                           Sts_FilterExcludedNumEvents => #instEventSortFilter_Alarm.Sts_FilterExcludedNumEvents,
                           Sts_SortFilterNumEvents => #instEventSortFilter_Alarm.Sts_SortFilterNumEvents);
END_REGION

REGION Network 10: *** Beging the WARNING area ****
END_REGION

REGION Network 11: Warning Event Summary Logic - Beginning Block
   // **********  WARNING SUMMATION  **********
   //  
   // The event summation begin instruction prepares the summation blocks.  It should be run each time before the FB_EventSummation blocks.
   RUNG wire#powerrail
      #instEventSumBeg_Warning(Sts_EventSummation := "Warning".Summation)
   END_RUNG
   // the same network as SCL:
   #instEventSumBeg_Warning(Sts_EventSummation := "Warning".Summation);   // "CPG_EventSummationBegin"
END_REGION

REGION Network 12: Warning Event Summary Logic - Unit Level Warnings
   RUNG wire#powerrail
      Contact( "UN".PackML_Sts.moduleActive )
      I_Contact( "HMI_Data".EMSortDisableWarning.Unit )
      #instEventSum_Warning_UN(In_EventStatus := "UN".Warning, Sts_EventSummation := "Warning".Summation, Sts_NumEvents => #instEventSum_Warning_UN.Sts_NumEvents, Sts_Category_0_Latched =>, Sts_Category_1_Latched =>, Sts_Category_2_Latched =>, Sts_Category_3_Latched =>, Sts_Category_4_Latched =>, Sts_Category_5_Latched =>, Sts_Category_6_Latched =>, Sts_Category_7_Latched =>, Sts_Category_8_Latched =>, Sts_Category_9_Latched =>, Sts_Category_0_NotLatched =>, Sts_Category_1_NotLatched =>, Sts_Category_2_NotLatched =>, Sts_Category_3_NotLatched =>, Sts_Category_4_NotLatched =>, Sts_Category_5_NotLatched =>, Sts_Category_6_NotLatched =>, Sts_Category_7_NotLatched =>, Sts_Category_8_NotLatched =>, Sts_Category_9_NotLatched =>, Sts_CurrentActiveEvent => #instEventSum_Warning_UN.Sts_CurrentActiveEvent, Sts_Error => #instEventSum_Warning_UN.Sts_Error, Sts_ErrorCode => #instEventSum_Warning_UN.Sts_ErrorCode)
   END_RUNG
   // the same network as SCL:
   IF "UN".PackML_Sts.moduleActive AND NOT "HMI_Data".EMSortDisableWarning.Unit THEN
       #instEventSum_Warning_UN(In_EventStatus := "UN".Warning,   // "CPG_EventSummation"
                               Sts_EventSummation := "Warning".Summation,
                               Sts_NumEvents => #instEventSum_Warning_UN.Sts_NumEvents,
                               Sts_CurrentActiveEvent => #instEventSum_Warning_UN.Sts_CurrentActiveEvent,
                               Sts_Error => #instEventSum_Warning_UN.Sts_Error,
                               Sts_ErrorCode => #instEventSum_Warning_UN.Sts_ErrorCode);
   END_IF;
END_REGION

REGION Network 13: Warning Event Summary Logic - Equipment Module #00
   // This instance of the Event Sum (or Event Summation) is used to merge the events 
   // from EM0 into the larger Unit or UN evevts list.
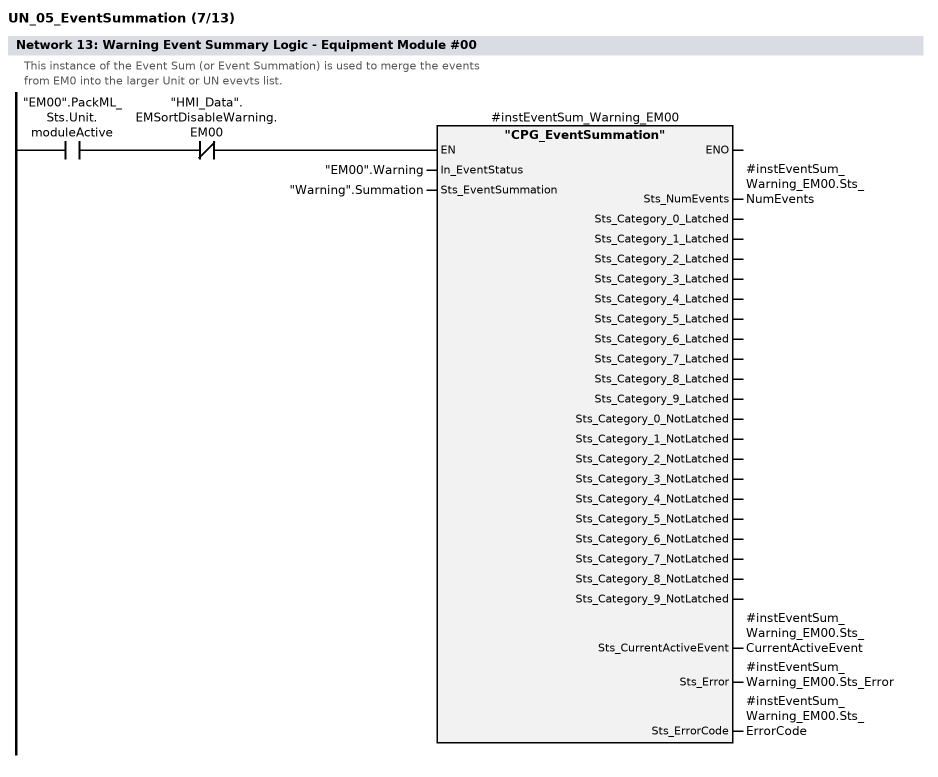
   RUNG wire#powerrail
      Contact( "EM00".PackML_Sts.Unit.moduleActive )
      I_Contact( "HMI_Data".EMSortDisableWarning.EM00 )
      #instEventSum_Warning_EM00(In_EventStatus := "EM00".Warning, Sts_EventSummation := "Warning".Summation, Sts_NumEvents => #instEventSum_Warning_EM00.Sts_NumEvents, Sts_Category_0_Latched =>, Sts_Category_1_Latched =>, Sts_Category_2_Latched =>, Sts_Category_3_Latched =>, Sts_Category_4_Latched =>, Sts_Category_5_Latched =>, Sts_Category_6_Latched =>, Sts_Category_7_Latched =>, Sts_Category_8_Latched =>, Sts_Category_9_Latched =>, Sts_Category_0_NotLatched =>, Sts_Category_1_NotLatched =>, Sts_Category_2_NotLatched =>, Sts_Category_3_NotLatched =>, Sts_Category_4_NotLatched =>, Sts_Category_5_NotLatched =>, Sts_Category_6_NotLatched =>, Sts_Category_7_NotLatched =>, Sts_Category_8_NotLatched =>, Sts_Category_9_NotLatched =>, Sts_CurrentActiveEvent => #instEventSum_Warning_EM00.Sts_CurrentActiveEvent, Sts_Error => #instEventSum_Warning_EM00.Sts_Error, Sts_ErrorCode => #instEventSum_Warning_EM00.Sts_ErrorCode)
   END_RUNG
   // the same network as SCL:
   IF "EM00".PackML_Sts.Unit.moduleActive AND NOT "HMI_Data".EMSortDisableWarning.EM00 THEN
       #instEventSum_Warning_EM00(In_EventStatus := "EM00".Warning,   // "CPG_EventSummation"
                               Sts_EventSummation := "Warning".Summation,
                               Sts_NumEvents => #instEventSum_Warning_EM00.Sts_NumEvents,
                               Sts_CurrentActiveEvent => #instEventSum_Warning_EM00.Sts_CurrentActiveEvent,
                               Sts_Error => #instEventSum_Warning_EM00.Sts_Error,
                               Sts_ErrorCode => #instEventSum_Warning_EM00.Sts_ErrorCode);
   END_IF;
END_REGION

REGION Network 14: Warning Event Summary Logic - Equipment Module #01
   // This instance of the Event Sum (or Event Summation) is used to merge the events 
   // from EM1 into the larger Unit or UN evevts list.
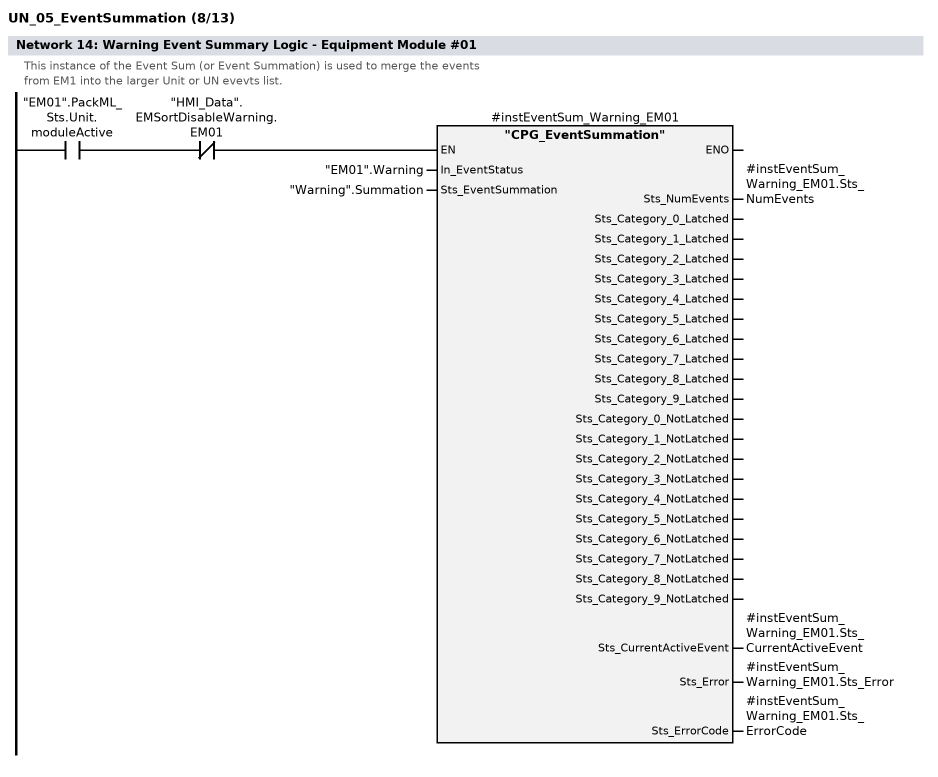
   RUNG wire#powerrail
      Contact( "EM01".PackML_Sts.Unit.moduleActive )
      I_Contact( "HMI_Data".EMSortDisableWarning.EM01 )
      #instEventSum_Warning_EM01(In_EventStatus := "EM01".Warning, Sts_EventSummation := "Warning".Summation, Sts_NumEvents => #instEventSum_Warning_EM01.Sts_NumEvents, Sts_Category_0_Latched =>, Sts_Category_1_Latched =>, Sts_Category_2_Latched =>, Sts_Category_3_Latched =>, Sts_Category_4_Latched =>, Sts_Category_5_Latched =>, Sts_Category_6_Latched =>, Sts_Category_7_Latched =>, Sts_Category_8_Latched =>, Sts_Category_9_Latched =>, Sts_Category_0_NotLatched =>, Sts_Category_1_NotLatched =>, Sts_Category_2_NotLatched =>, Sts_Category_3_NotLatched =>, Sts_Category_4_NotLatched =>, Sts_Category_5_NotLatched =>, Sts_Category_6_NotLatched =>, Sts_Category_7_NotLatched =>, Sts_Category_8_NotLatched =>, Sts_Category_9_NotLatched =>, Sts_CurrentActiveEvent => #instEventSum_Warning_EM01.Sts_CurrentActiveEvent, Sts_Error => #instEventSum_Warning_EM01.Sts_Error, Sts_ErrorCode => #instEventSum_Warning_EM01.Sts_ErrorCode)
   END_RUNG
   // the same network as SCL:
   IF "EM01".PackML_Sts.Unit.moduleActive AND NOT "HMI_Data".EMSortDisableWarning.EM01 THEN
       #instEventSum_Warning_EM01(In_EventStatus := "EM01".Warning,   // "CPG_EventSummation"
                               Sts_EventSummation := "Warning".Summation,
                               Sts_NumEvents => #instEventSum_Warning_EM01.Sts_NumEvents,
                               Sts_CurrentActiveEvent => #instEventSum_Warning_EM01.Sts_CurrentActiveEvent,
                               Sts_Error => #instEventSum_Warning_EM01.Sts_Error,
                               Sts_ErrorCode => #instEventSum_Warning_EM01.Sts_ErrorCode);
   END_IF;
END_REGION

REGION Network 15: Warning Event Summary Logic - Equipment Module #02
   // This instance of the Event Sum (or Event Summation) is used to merge the events 
   // from EM01 into the larger Unit or UN evevts list.
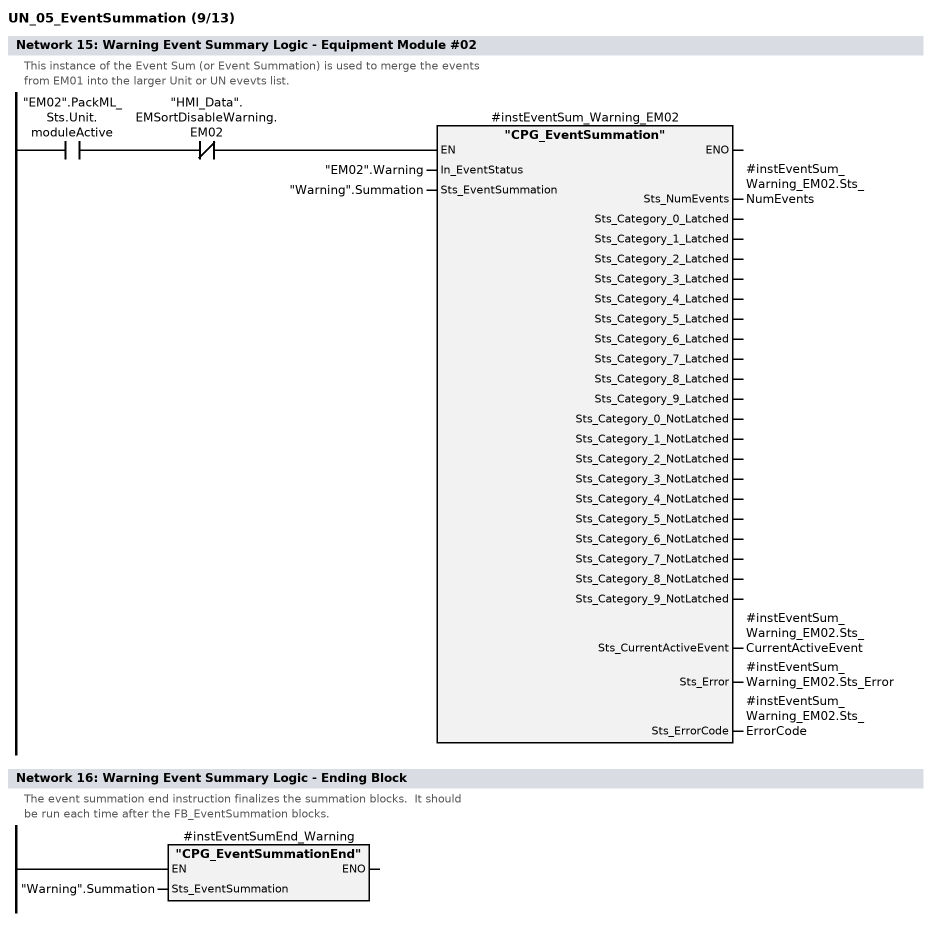
   RUNG wire#powerrail
      Contact( "EM02".PackML_Sts.Unit.moduleActive )
      I_Contact( "HMI_Data".EMSortDisableWarning.EM02 )
      #instEventSum_Warning_EM02(In_EventStatus := "EM02".Warning, Sts_EventSummation := "Warning".Summation, Sts_NumEvents => #instEventSum_Warning_EM02.Sts_NumEvents, Sts_Category_0_Latched =>, Sts_Category_1_Latched =>, Sts_Category_2_Latched =>, Sts_Category_3_Latched =>, Sts_Category_4_Latched =>, Sts_Category_5_Latched =>, Sts_Category_6_Latched =>, Sts_Category_7_Latched =>, Sts_Category_8_Latched =>, Sts_Category_9_Latched =>, Sts_Category_0_NotLatched =>, Sts_Category_1_NotLatched =>, Sts_Category_2_NotLatched =>, Sts_Category_3_NotLatched =>, Sts_Category_4_NotLatched =>, Sts_Category_5_NotLatched =>, Sts_Category_6_NotLatched =>, Sts_Category_7_NotLatched =>, Sts_Category_8_NotLatched =>, Sts_Category_9_NotLatched =>, Sts_CurrentActiveEvent => #instEventSum_Warning_EM02.Sts_CurrentActiveEvent, Sts_Error => #instEventSum_Warning_EM02.Sts_Error, Sts_ErrorCode => #instEventSum_Warning_EM02.Sts_ErrorCode)
   END_RUNG
   // the same network as SCL:
   IF "EM02".PackML_Sts.Unit.moduleActive AND NOT "HMI_Data".EMSortDisableWarning.EM02 THEN
       #instEventSum_Warning_EM02(In_EventStatus := "EM02".Warning,   // "CPG_EventSummation"
                               Sts_EventSummation := "Warning".Summation,
                               Sts_NumEvents => #instEventSum_Warning_EM02.Sts_NumEvents,
                               Sts_CurrentActiveEvent => #instEventSum_Warning_EM02.Sts_CurrentActiveEvent,
                               Sts_Error => #instEventSum_Warning_EM02.Sts_Error,
                               Sts_ErrorCode => #instEventSum_Warning_EM02.Sts_ErrorCode);
   END_IF;
END_REGION

REGION Network 16: Warning Event Summary Logic - Ending Block
   // The event summation end instruction finalizes the summation blocks.  It should 
   // be run each time after the FB_EventSummation blocks.
   RUNG wire#powerrail
      #instEventSumEnd_Warning(Sts_EventSummation := "Warning".Summation)
   END_RUNG
   // the same network as SCL:
   #instEventSumEnd_Warning(Sts_EventSummation := "Warning".Summation);   // "CPG_EventSummationEnd"
END_REGION

REGION Network 17: Event Sort Filter logic - Warnings
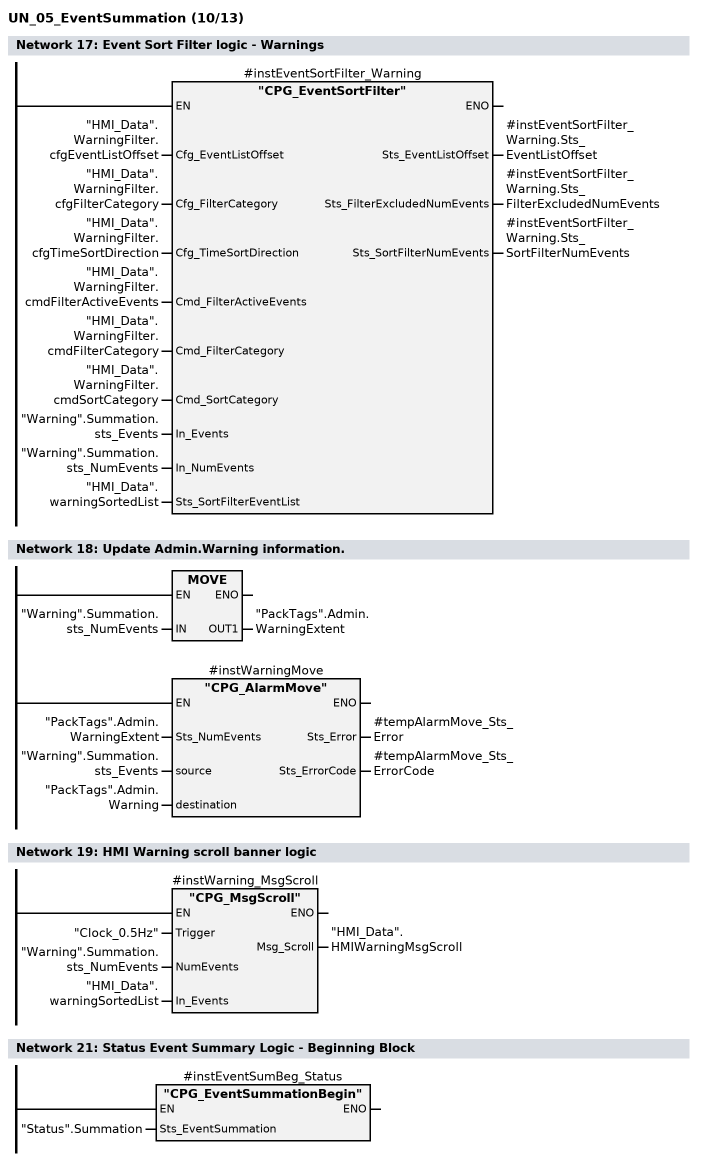
   RUNG wire#powerrail
      #instEventSortFilter_Warning(Cfg_EventListOffset := "HMI_Data".WarningFilter.cfgEventListOffset, Cfg_FilterCategory := "HMI_Data".WarningFilter.cfgFilterCategory, Cfg_TimeSortDirection := "HMI_Data".WarningFilter.cfgTimeSortDirection, Cmd_FilterActiveEvents := "HMI_Data".WarningFilter.cmdFilterActiveEvents, Cmd_FilterCategory := "HMI_Data".WarningFilter.cmdFilterCategory, Cmd_SortCategory := "HMI_Data".WarningFilter.cmdSortCategory, In_Events := "Warning".Summation.sts_Events, In_NumEvents := "Warning".Summation.sts_NumEvents, Sts_SortFilterEventList := "HMI_Data".warningSortedList, Sts_EventListOffset => #instEventSortFilter_Warning.Sts_EventListOffset, Sts_FilterExcludedNumEvents => #instEventSortFilter_Warning.Sts_FilterExcludedNumEvents, Sts_SortFilterNumEvents => #instEventSortFilter_Warning.Sts_SortFilterNumEvents)
   END_RUNG
   // the same network as SCL:
   #instEventSortFilter_Warning(Cfg_EventListOffset := "HMI_Data".WarningFilter.cfgEventListOffset,   // "CPG_EventSortFilter"
                           Cfg_FilterCategory := "HMI_Data".WarningFilter.cfgFilterCategory,
                           Cfg_TimeSortDirection := "HMI_Data".WarningFilter.cfgTimeSortDirection,
                           Cmd_FilterActiveEvents := "HMI_Data".WarningFilter.cmdFilterActiveEvents,
                           Cmd_FilterCategory := "HMI_Data".WarningFilter.cmdFilterCategory,
                           Cmd_SortCategory := "HMI_Data".WarningFilter.cmdSortCategory,
                           In_Events := "Warning".Summation.sts_Events,
                           In_NumEvents := "Warning".Summation.sts_NumEvents,
                           Sts_SortFilterEventList := "HMI_Data".warningSortedList,
                           Sts_EventListOffset => #instEventSortFilter_Warning.Sts_EventListOffset,
                           Sts_FilterExcludedNumEvents => #instEventSortFilter_Warning.Sts_FilterExcludedNumEvents,
                           Sts_SortFilterNumEvents => #instEventSortFilter_Warning.Sts_SortFilterNumEvents);
END_REGION

REGION Network 18: Update Admin.Warning information.
   RUNG wire#powerrail
      { S7_GenerateENO := "TRUE" } Move(in := "Warning".Summation.sts_NumEvents, out1 => "PackTags".Admin.WarningExtent)
   END_RUNG
   RUNG wire#powerrail
      #instWarningMove(Sts_NumEvents := "PackTags".Admin.WarningExtent, source := "Warning".Summation.sts_Events, destination := "PackTags".Admin.Warning, Sts_Error => #tempAlarmMove_Sts_Error, Sts_ErrorCode => #tempAlarmMove_Sts_ErrorCode)
   END_RUNG
   // the same network as SCL:
   "PackTags".Admin.WarningExtent := "Warning".Summation.sts_NumEvents;
   #instWarningMove(Sts_NumEvents := "PackTags".Admin.WarningExtent,   // "CPG_AlarmMove"
                    source := "Warning".Summation.sts_Events,
                    destination := "PackTags".Admin.Warning,
                    Sts_Error => #tempAlarmMove_Sts_Error,
                    Sts_ErrorCode => #tempAlarmMove_Sts_ErrorCode);
END_REGION

REGION Network 19: HMI Warning scroll banner logic
   RUNG wire#powerrail
      #instWarning_MsgScroll(Trigger := "Clock_0.5Hz", NumEvents := "Warning".Summation.sts_NumEvents, In_Events := "HMI_Data".warningSortedList, Msg_Scroll => "HMI_Data".HMIWarningMsgScroll)
   END_RUNG
   // the same network as SCL:
   #instWarning_MsgScroll(Trigger := "Clock_0.5Hz",   // "CPG_MsgScroll"
                          NumEvents := "Warning".Summation.sts_NumEvents,
                          In_Events := "HMI_Data".warningSortedList,
                          Msg_Scroll => "HMI_Data".HMIWarningMsgScroll);
END_REGION

REGION Network 20: *** Status Event Summation ***
END_REGION

REGION Network 21: Status Event Summary Logic - Beginning Block
   RUNG wire#powerrail
      #instEventSumBeg_Status(Sts_EventSummation := "Status".Summation)
   END_RUNG
   // the same network as SCL:
   #instEventSumBeg_Status(Sts_EventSummation := "Status".Summation);   // "CPG_EventSummationBegin"
END_REGION

REGION Network 22: Status Event Summary Logic - Unit
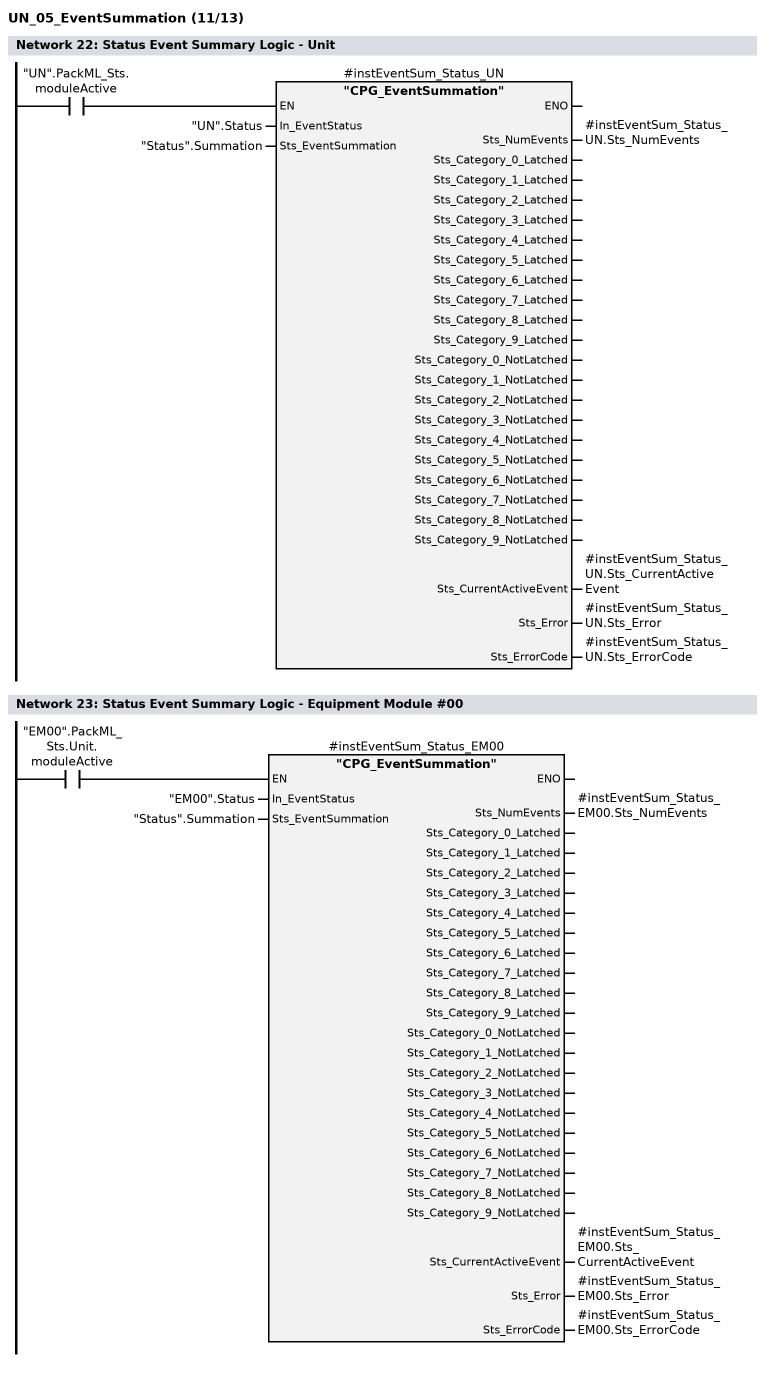
   RUNG wire#powerrail
      Contact( "UN".PackML_Sts.moduleActive )
      #instEventSum_Status_UN(In_EventStatus := "UN".Status, Sts_EventSummation := "Status".Summation, Sts_NumEvents => #instEventSum_Status_UN.Sts_NumEvents, Sts_Category_0_Latched =>, Sts_Category_1_Latched =>, Sts_Category_2_Latched =>, Sts_Category_3_Latched =>, Sts_Category_4_Latched =>, Sts_Category_5_Latched =>, Sts_Category_6_Latched =>, Sts_Category_7_Latched =>, Sts_Category_8_Latched =>, Sts_Category_9_Latched =>, Sts_Category_0_NotLatched =>, Sts_Category_1_NotLatched =>, Sts_Category_2_NotLatched =>, Sts_Category_3_NotLatched =>, Sts_Category_4_NotLatched =>, Sts_Category_5_NotLatched =>, Sts_Category_6_NotLatched =>, Sts_Category_7_NotLatched =>, Sts_Category_8_NotLatched =>, Sts_Category_9_NotLatched =>, Sts_CurrentActiveEvent => #instEventSum_Status_UN.Sts_CurrentActiveEvent, Sts_Error => #instEventSum_Status_UN.Sts_Error, Sts_ErrorCode => #instEventSum_Status_UN.Sts_ErrorCode)
   END_RUNG
   // the same network as SCL:
   IF "UN".PackML_Sts.moduleActive THEN
       #instEventSum_Status_UN(In_EventStatus := "UN".Status,   // "CPG_EventSummation"
                               Sts_EventSummation := "Status".Summation,
                               Sts_NumEvents => #instEventSum_Status_UN.Sts_NumEvents,
                               Sts_CurrentActiveEvent => #instEventSum_Status_UN.Sts_CurrentActiveEvent,
                               Sts_Error => #instEventSum_Status_UN.Sts_Error,
                               Sts_ErrorCode => #instEventSum_Status_UN.Sts_ErrorCode);
   END_IF;
END_REGION

REGION Network 23: Status Event Summary Logic - Equipment Module #00
   RUNG wire#powerrail
      Contact( "EM00".PackML_Sts.Unit.moduleActive )
      #instEventSum_Status_EM00(In_EventStatus := "EM00".Status, Sts_EventSummation := "Status".Summation, Sts_NumEvents => #instEventSum_Status_EM00.Sts_NumEvents, Sts_Category_0_Latched =>, Sts_Category_1_Latched =>, Sts_Category_2_Latched =>, Sts_Category_3_Latched =>, Sts_Category_4_Latched =>, Sts_Category_5_Latched =>, Sts_Category_6_Latched =>, Sts_Category_7_Latched =>, Sts_Category_8_Latched =>, Sts_Category_9_Latched =>, Sts_Category_0_NotLatched =>, Sts_Category_1_NotLatched =>, Sts_Category_2_NotLatched =>, Sts_Category_3_NotLatched =>, Sts_Category_4_NotLatched =>, Sts_Category_5_NotLatched =>, Sts_Category_6_NotLatched =>, Sts_Category_7_NotLatched =>, Sts_Category_8_NotLatched =>, Sts_Category_9_NotLatched =>, Sts_CurrentActiveEvent => #instEventSum_Status_EM00.Sts_CurrentActiveEvent, Sts_Error => #instEventSum_Status_EM00.Sts_Error, Sts_ErrorCode => #instEventSum_Status_EM00.Sts_ErrorCode)
   END_RUNG
   // the same network as SCL:
   IF "EM00".PackML_Sts.Unit.moduleActive THEN
       #instEventSum_Status_EM00(In_EventStatus := "EM00".Status,   // "CPG_EventSummation"
                               Sts_EventSummation := "Status".Summation,
                               Sts_NumEvents => #instEventSum_Status_EM00.Sts_NumEvents,
                               Sts_CurrentActiveEvent => #instEventSum_Status_EM00.Sts_CurrentActiveEvent,
                               Sts_Error => #instEventSum_Status_EM00.Sts_Error,
                               Sts_ErrorCode => #instEventSum_Status_EM00.Sts_ErrorCode);
   END_IF;
END_REGION

REGION Network 24: Status Event Summary Logic - Equipment Module #01
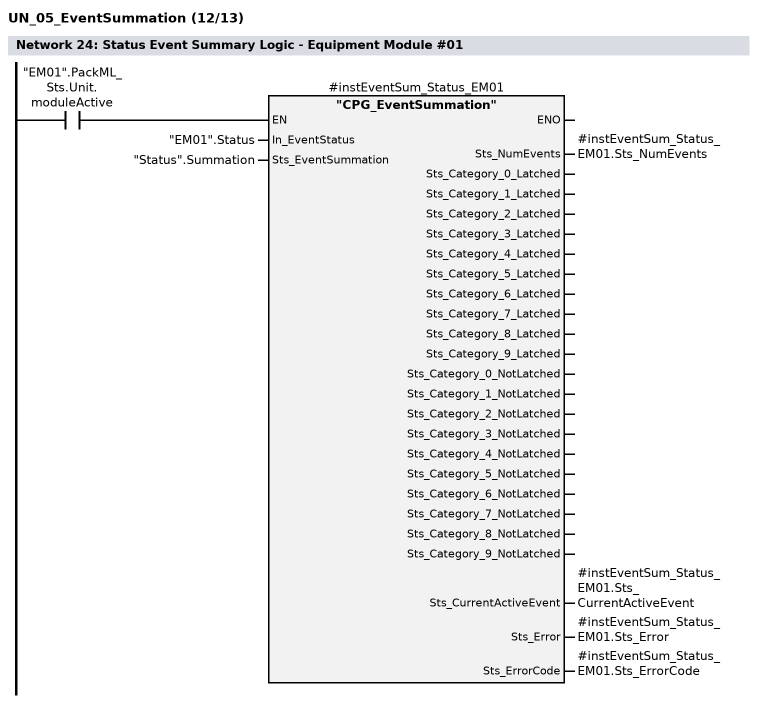
   RUNG wire#powerrail
      Contact( "EM01".PackML_Sts.Unit.moduleActive )
      #instEventSum_Status_EM01(In_EventStatus := "EM01".Status, Sts_EventSummation := "Status".Summation, Sts_NumEvents => #instEventSum_Status_EM01.Sts_NumEvents, Sts_Category_0_Latched =>, Sts_Category_1_Latched =>, Sts_Category_2_Latched =>, Sts_Category_3_Latched =>, Sts_Category_4_Latched =>, Sts_Category_5_Latched =>, Sts_Category_6_Latched =>, Sts_Category_7_Latched =>, Sts_Category_8_Latched =>, Sts_Category_9_Latched =>, Sts_Category_0_NotLatched =>, Sts_Category_1_NotLatched =>, Sts_Category_2_NotLatched =>, Sts_Category_3_NotLatched =>, Sts_Category_4_NotLatched =>, Sts_Category_5_NotLatched =>, Sts_Category_6_NotLatched =>, Sts_Category_7_NotLatched =>, Sts_Category_8_NotLatched =>, Sts_Category_9_NotLatched =>, Sts_CurrentActiveEvent => #instEventSum_Status_EM01.Sts_CurrentActiveEvent, Sts_Error => #instEventSum_Status_EM01.Sts_Error, Sts_ErrorCode => #instEventSum_Status_EM01.Sts_ErrorCode)
   END_RUNG
   // the same network as SCL:
   IF "EM01".PackML_Sts.Unit.moduleActive THEN
       #instEventSum_Status_EM01(In_EventStatus := "EM01".Status,   // "CPG_EventSummation"
                               Sts_EventSummation := "Status".Summation,
                               Sts_NumEvents => #instEventSum_Status_EM01.Sts_NumEvents,
                               Sts_CurrentActiveEvent => #instEventSum_Status_EM01.Sts_CurrentActiveEvent,
                               Sts_Error => #instEventSum_Status_EM01.Sts_Error,
                               Sts_ErrorCode => #instEventSum_Status_EM01.Sts_ErrorCode);
   END_IF;
END_REGION

REGION Network 25: Status Event Summary Logic - Equipment Module #02
   // This instance of the Event Sum (or Event Summation) is used to merge the events 
   // from EM01 into the larger Unit or UN evevts list.
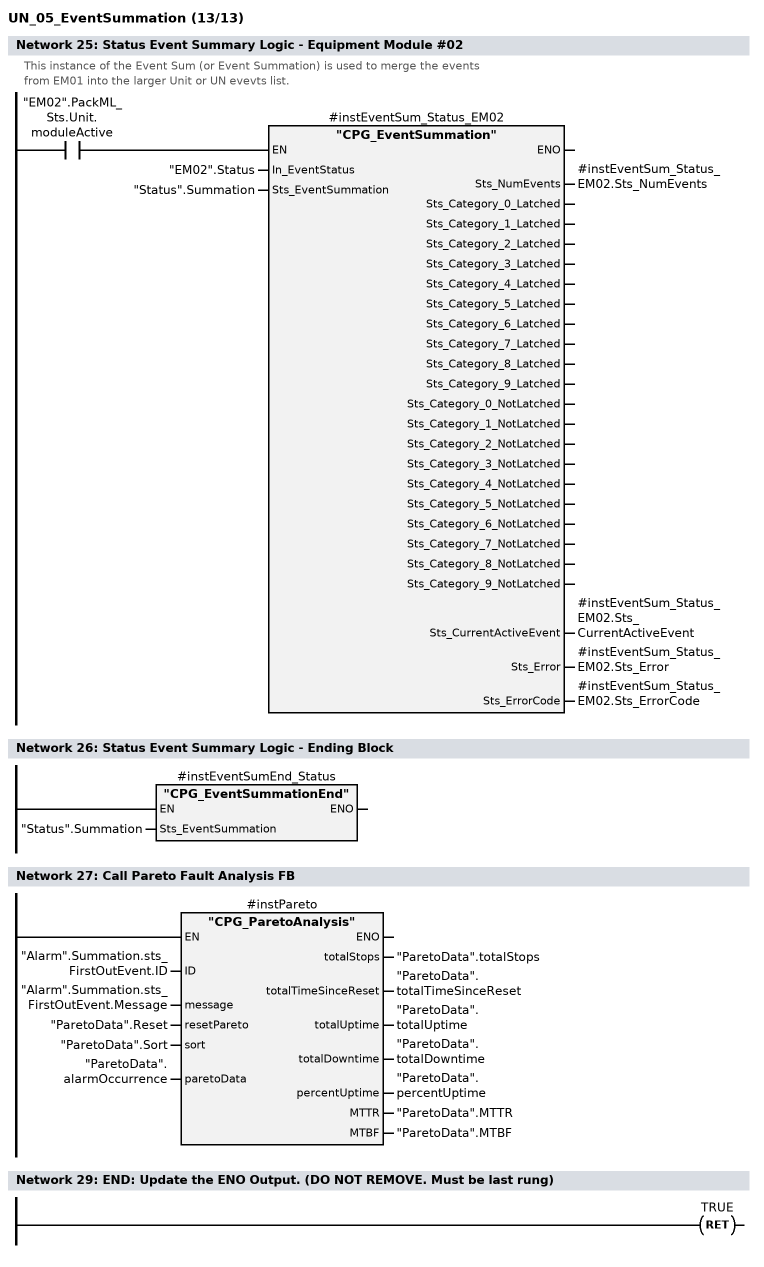
   RUNG wire#powerrail
      Contact( "EM02".PackML_Sts.Unit.moduleActive )
      #instEventSum_Status_EM02(In_EventStatus := "EM02".Status, Sts_EventSummation := "Status".Summation, Sts_NumEvents => #instEventSum_Status_EM02.Sts_NumEvents, Sts_Category_0_Latched =>, Sts_Category_1_Latched =>, Sts_Category_2_Latched =>, Sts_Category_3_Latched =>, Sts_Category_4_Latched =>, Sts_Category_5_Latched =>, Sts_Category_6_Latched =>, Sts_Category_7_Latched =>, Sts_Category_8_Latched =>, Sts_Category_9_Latched =>, Sts_Category_0_NotLatched =>, Sts_Category_1_NotLatched =>, Sts_Category_2_NotLatched =>, Sts_Category_3_NotLatched =>, Sts_Category_4_NotLatched =>, Sts_Category_5_NotLatched =>, Sts_Category_6_NotLatched =>, Sts_Category_7_NotLatched =>, Sts_Category_8_NotLatched =>, Sts_Category_9_NotLatched =>, Sts_CurrentActiveEvent => #instEventSum_Status_EM02.Sts_CurrentActiveEvent, Sts_Error => #instEventSum_Status_EM02.Sts_Error, Sts_ErrorCode => #instEventSum_Status_EM02.Sts_ErrorCode)
   END_RUNG
   // the same network as SCL:
   IF "EM02".PackML_Sts.Unit.moduleActive THEN
       #instEventSum_Status_EM02(In_EventStatus := "EM02".Status,   // "CPG_EventSummation"
                               Sts_EventSummation := "Status".Summation,
                               Sts_NumEvents => #instEventSum_Status_EM02.Sts_NumEvents,
                               Sts_CurrentActiveEvent => #instEventSum_Status_EM02.Sts_CurrentActiveEvent,
                               Sts_Error => #instEventSum_Status_EM02.Sts_Error,
                               Sts_ErrorCode => #instEventSum_Status_EM02.Sts_ErrorCode);
   END_IF;
END_REGION

REGION Network 26: Status Event Summary Logic - Ending Block
   RUNG wire#powerrail
      #instEventSumEnd_Status(Sts_EventSummation := "Status".Summation)
   END_RUNG
   // the same network as SCL:
   #instEventSumEnd_Status(Sts_EventSummation := "Status".Summation);   // "CPG_EventSummationEnd"
END_REGION

REGION Network 27: Call Pareto Fault Analysis FB
   RUNG wire#powerrail
      #instPareto(ID := "Alarm".Summation.sts_FirstOutEvent.ID, message := "Alarm".Summation.sts_FirstOutEvent.Message, resetPareto := "ParetoData".Reset, sort := "ParetoData".Sort, paretoData := "ParetoData".alarmOccurrence, totalStops => "ParetoData".totalStops, totalTimeSinceReset => "ParetoData".totalTimeSinceReset, totalUptime => "ParetoData".totalUptime, totalDowntime => "ParetoData".totalDowntime, percentUptime => "ParetoData".percentUptime, MTTR => "ParetoData".MTTR, MTBF => "ParetoData".MTBF)
   END_RUNG
   // the same network as SCL:
   #instPareto(ID := "Alarm".Summation.sts_FirstOutEvent.ID,   // "CPG_ParetoAnalysis"
               message := "Alarm".Summation.sts_FirstOutEvent.Message,
               resetPareto := "ParetoData".Reset,
               sort := "ParetoData".Sort,
               paretoData := "ParetoData".alarmOccurrence,
               totalStops => "ParetoData".totalStops,
               totalTimeSinceReset => "ParetoData".totalTimeSinceReset,
               totalUptime => "ParetoData".totalUptime,
               totalDowntime => "ParetoData".totalDowntime,
               percentUptime => "ParetoData".percentUptime,
               MTTR => "ParetoData".MTTR,
               MTBF => "ParetoData".MTBF);
END_REGION

REGION Network 28: HMI Warning scroll banner logic
END_REGION

REGION Network 29: END: Update the ENO Output. (DO NOT REMOVE. Must be last rung)
   RUNG wire#powerrail
      ReturnCoil( TRUE )
   END_RUNG
   // the same network as SCL:
   ENO := TRUE;
   RETURN;
END_REGION
END_FUNCTION_BLOCK

FUNCTION_BLOCK "UN_06_MiscFunctions"   // FB31626, LAD
TITLE = UN_06_MiscFunctions
{ S7_Optimized_Access := 'TRUE' }
AUTHOR : tech.team.motioncontrol@siemens.com
FAMILY : CPG
VERSION : 1.1
// Support: tech.team.motioncontrol@siemens.com
   VAR
      instOEE_Calculation : "CPG_OEE";   // FB used to calculate the real-time OEE value
      statOneShot_ProdConsumerCounter : Bool;   // One Shot - products consumed counter
      statOneShot_ProdProcessedCounter : Bool;   // One Shot - products processed counter
      statOneShot_ProdDefectiveCounter : Bool;   // One Shot - products defective counter
   END_VAR
   VAR_TEMP
      tempReadClockRetVal : Int;
      tempProductionCounterTrigger : Bool;
   END_VAR
   VAR_TEMP   // added for the SCL form of the ladder/FBD networks
      _w1 : Bool;
   END_VAR
BEGIN

REGION Network 1: Update the PackTags Admin.PLC_Date_Time with current PLC time
   // 1) Update the "PackTags".Admin.PLC_Date_Time with the current PLC time.
   // 2) Update "HMI_Data".PLC_Date_Time.DATE_TIME with current PLC time so the HMI 
   // and PLC are time synchronized.
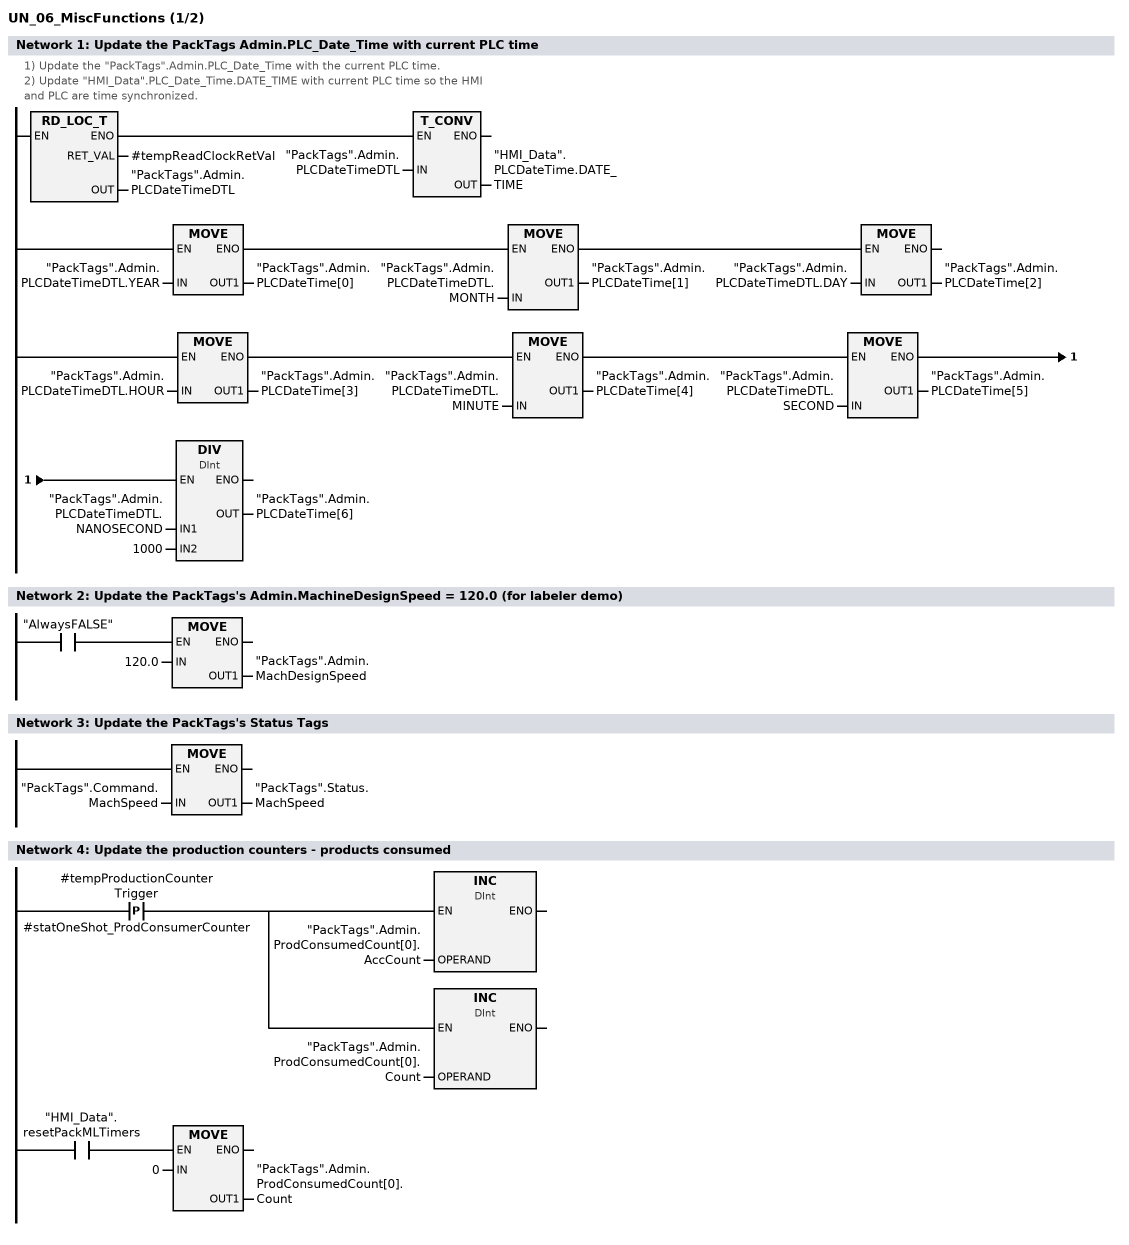
   // ENO of a box is taken as its EN; it also drops when the box reports an error
   #tempReadClockRetVal := RD_LOC_T(OUT => "PackTags".Admin.PLCDateTimeDTL);
   "HMI_Data".PLCDateTime.DATE_TIME := T_CONV(IN := "PackTags".Admin.PLCDateTimeDTL);
   "PackTags".Admin.PLCDateTime[0] := "PackTags".Admin.PLCDateTimeDTL.YEAR;
   "PackTags".Admin.PLCDateTime[1] := "PackTags".Admin.PLCDateTimeDTL.MONTH;
   "PackTags".Admin.PLCDateTime[2] := "PackTags".Admin.PLCDateTimeDTL.DAY;
   "PackTags".Admin.PLCDateTime[3] := "PackTags".Admin.PLCDateTimeDTL.HOUR;
   "PackTags".Admin.PLCDateTime[4] := "PackTags".Admin.PLCDateTimeDTL.MINUTE;
   "PackTags".Admin.PLCDateTime[5] := "PackTags".Admin.PLCDateTimeDTL.SECOND;
   "PackTags".Admin.PLCDateTime[6] := "PackTags".Admin.PLCDateTimeDTL.NANOSECOND / 1000;
END_REGION

REGION Network 2: Update the PackTags's Admin.MachineDesignSpeed = 120.0 (for labeler demo)
   RUNG wire#powerrail
      Contact( "AlwaysFALSE" )
      Move(in := 120.0, out1 => "PackTags".Admin.MachDesignSpeed)
   END_RUNG
   // the same network as SCL:
   IF "AlwaysFALSE" THEN "PackTags".Admin.MachDesignSpeed := 120.0; END_IF;
END_REGION

REGION Network 3: Update the PackTags's Status Tags
   RUNG wire#powerrail
      Move(in := "PackTags".Command.MachSpeed, out1 => "PackTags".Status.MachSpeed)
   END_RUNG
   // the same network as SCL:
   "PackTags".Status.MachSpeed := "PackTags".Command.MachSpeed;
END_REGION

REGION Network 4: Update the production counters - products consumed
   RUNG wire#powerrail
      P_Contact(operand := #tempProductionCounterTrigger, bit := #statOneShot_ProdConsumerCounter)
      wire#w1
      { S7_Templates := "DestType := DInt" } Inc( "PackTags".Admin.ProdConsumedCount[0].AccCount )
   END_RUNG
   RUNG wire#w1
      { S7_Templates := "DestType := DInt" } Inc( "PackTags".Admin.ProdConsumedCount[0].Count )
   END_RUNG
   RUNG wire#powerrail
      Contact( "HMI_Data".resetPackMLTimers )
      Move(in := 0, out1 => "PackTags".Admin.ProdConsumedCount[0].Count)
   END_RUNG
   // the same network as SCL:
   #_w1 := #tempProductionCounterTrigger AND NOT #statOneShot_ProdConsumerCounter;   // rising edge of #tempProductionCounterTrigger
   #statOneShot_ProdConsumerCounter := #tempProductionCounterTrigger;
   IF #_w1 THEN
       "PackTags".Admin.ProdConsumedCount[0].AccCount := "PackTags".Admin.ProdConsumedCount[0].AccCount + 1;
       "PackTags".Admin.ProdConsumedCount[0].Count := "PackTags".Admin.ProdConsumedCount[0].Count + 1;
   END_IF;
   IF "HMI_Data".resetPackMLTimers THEN "PackTags".Admin.ProdConsumedCount[0].Count := 0; END_IF;
END_REGION

REGION Network 5: Update the production counters - products processed
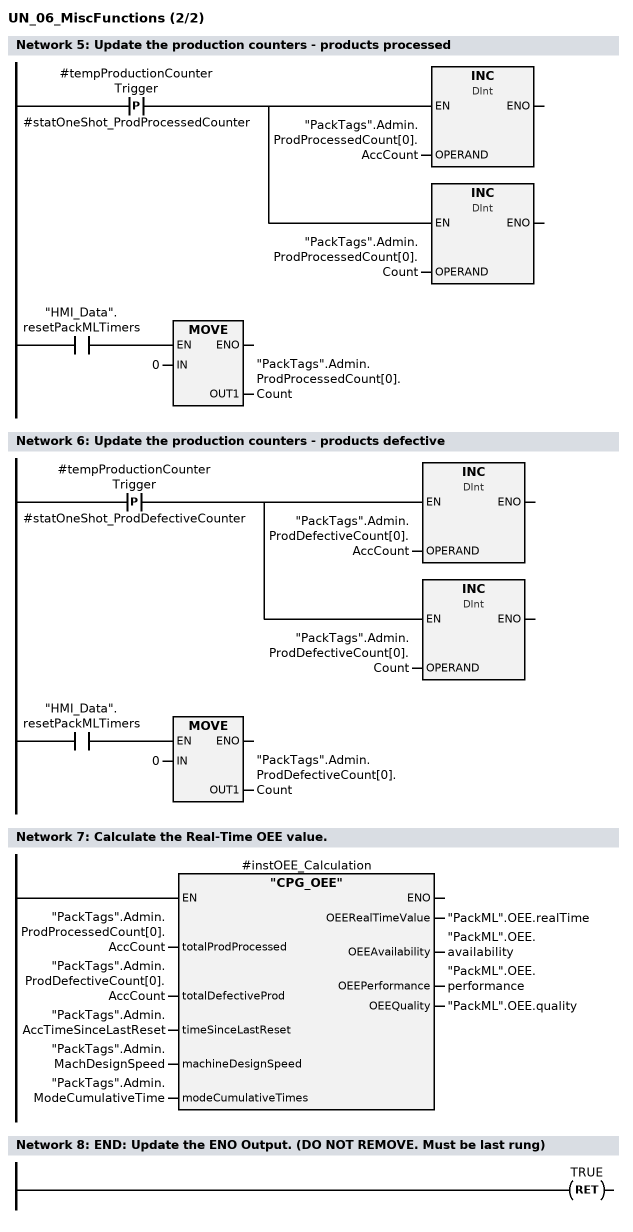
   RUNG wire#powerrail
      P_Contact(operand := #tempProductionCounterTrigger, bit := #statOneShot_ProdProcessedCounter)
      wire#w1
      { S7_Templates := "DestType := DInt" } Inc( "PackTags".Admin.ProdProcessedCount[0].AccCount )
   END_RUNG
   RUNG wire#w1
      { S7_Templates := "DestType := DInt" } Inc( "PackTags".Admin.ProdProcessedCount[0].Count )
   END_RUNG
   RUNG wire#powerrail
      Contact( "HMI_Data".resetPackMLTimers )
      Move(in := 0, out1 => "PackTags".Admin.ProdProcessedCount[0].Count)
   END_RUNG
   // the same network as SCL:
   #_w1 := #tempProductionCounterTrigger AND NOT #statOneShot_ProdProcessedCounter;   // rising edge of #tempProductionCounterTrigger
   #statOneShot_ProdProcessedCounter := #tempProductionCounterTrigger;
   IF #_w1 THEN
       "PackTags".Admin.ProdProcessedCount[0].AccCount := "PackTags".Admin.ProdProcessedCount[0].AccCount + 1;
       "PackTags".Admin.ProdProcessedCount[0].Count := "PackTags".Admin.ProdProcessedCount[0].Count + 1;
   END_IF;
   IF "HMI_Data".resetPackMLTimers THEN "PackTags".Admin.ProdProcessedCount[0].Count := 0; END_IF;
END_REGION

REGION Network 6: Update the production counters - products defective
   RUNG wire#powerrail
      P_Contact(operand := #tempProductionCounterTrigger, bit := #statOneShot_ProdDefectiveCounter)
      wire#w1
      { S7_Templates := "DestType := DInt" } Inc( "PackTags".Admin.ProdDefectiveCount[0].AccCount )
   END_RUNG
   RUNG wire#w1
      { S7_Templates := "DestType := DInt" } Inc( "PackTags".Admin.ProdDefectiveCount[0].Count )
   END_RUNG
   RUNG wire#powerrail
      Contact( "HMI_Data".resetPackMLTimers )
      Move(in := 0, out1 => "PackTags".Admin.ProdDefectiveCount[0].Count)
   END_RUNG
   // the same network as SCL:
   #_w1 := #tempProductionCounterTrigger AND NOT #statOneShot_ProdDefectiveCounter;   // rising edge of #tempProductionCounterTrigger
   #statOneShot_ProdDefectiveCounter := #tempProductionCounterTrigger;
   IF #_w1 THEN
       "PackTags".Admin.ProdDefectiveCount[0].AccCount := "PackTags".Admin.ProdDefectiveCount[0].AccCount + 1;
       "PackTags".Admin.ProdDefectiveCount[0].Count := "PackTags".Admin.ProdDefectiveCount[0].Count + 1;
   END_IF;
   IF "HMI_Data".resetPackMLTimers THEN "PackTags".Admin.ProdDefectiveCount[0].Count := 0; END_IF;
END_REGION

REGION Network 7: Calculate the Real-Time OEE value.
   RUNG wire#powerrail
      #instOEE_Calculation(totalProdProcessed := "PackTags".Admin.ProdProcessedCount[0].AccCount, totalDefectiveProd := "PackTags".Admin.ProdDefectiveCount[0].AccCount, timeSinceLastReset := "PackTags".Admin.AccTimeSinceLastReset, machineDesignSpeed := "PackTags".Admin.MachDesignSpeed, modeCumulativeTimes := "PackTags".Admin.ModeCumulativeTime, OEERealTimeValue => "PackML".OEE.realTime, OEEAvailability => "PackML".OEE.availability, OEEPerformance => "PackML".OEE.performance, OEEQuality => "PackML".OEE.quality)
   END_RUNG
   // the same network as SCL:
   #instOEE_Calculation(totalProdProcessed := "PackTags".Admin.ProdProcessedCount[0].AccCount,   // "CPG_OEE"
                        totalDefectiveProd := "PackTags".Admin.ProdDefectiveCount[0].AccCount,
                        timeSinceLastReset := "PackTags".Admin.AccTimeSinceLastReset,
                        machineDesignSpeed := "PackTags".Admin.MachDesignSpeed,
                        modeCumulativeTimes := "PackTags".Admin.ModeCumulativeTime,
                        OEERealTimeValue => "PackML".OEE.realTime,
                        OEEAvailability => "PackML".OEE.availability,
                        OEEPerformance => "PackML".OEE.performance,
                        OEEQuality => "PackML".OEE.quality);
END_REGION
